FUNCTION_BLOCK "FB_ManInsp_V1.00"   // FB24, LAD
{ S7_Optimized_Access := 'TRUE' }
VERSION : 0.1
   VAR_INPUT
      IN_xCycleON : Bool;   // Cycle ON
      IN_xCycleONDel : Bool;   // Delayed cycle ON signal
      IN_xGeneralReset : Bool;   // General reset
      IN_xResetAlarms : Bool;   // Reset alarms
      IN_xFaultsEnabled : Bool;   // Faults enabled
      IN_dGlassBreakMachineIndex : DInt;   // Glass break machine index
      IN_dNumButtonDefect : DInt;   // Number of defect button
      IN_dNumQltDefect : DInt;   // Number of quality defect
      INPUT : Struct   // Digital inputs
         xPowerSupplyControl : Bool;   // L+.Power supply control
         xOpenRolls : Bool;   // SA.Open rolls
         xCloseRolls : Bool;   // SA.Close rolls
         rgxDefectButtons : Array[0..#CONST_MAX_DEFECT_BUTTONS_IND] of Bool;   // Defects buttons
         rgxQualityButtons : Array[0..#CONST_MAX_QUALITY_BUTTONS_IND] of Bool;   // Quality buttons
      END_STRUCT;
   END_VAR
   VAR_OUTPUT
      OUTPUT : Struct
         xFanCommand : Bool;   // Fan command
         xCloseRolls : Bool;   // YV.Close rolls
         xOpenRolls : Bool;   // YV.Open rolls
         xLampOpenCloseRolls : Bool;   // HL.Open/Close rolls
         rgxDefectButtonsLamp : Array[0..#CONST_MAX_DEFECT_BUTTONS_IND] of Bool;   // Defect buttons lamp
         rgxQualityButtonsLamp : Array[0..#CONST_MAX_QUALITY_BUTTONS_IND] of Bool;   // quality buttons lamp
      END_STRUCT;
   END_VAR
   VAR_IN_OUT
      INO_tFBAddDefect : "FB_Defects_Add_V1.00";   // Add defect DB
      INO_tOBInitialize : "GP_OB_Initialize";   // OB Initialize
      INO_tEncoder : "UDT_Encoder";   // Encoder data
      INO_tRibbon : "UDT_RibbonData";   // Ribbon data
      INO_xDefectBufferFull : Bool;   // Defect buffer full
   END_VAR
   VAR RETAIN
      tHMW : Struct   // HMI Write
         tMan : Struct   // Manual commands
            xFanCommand : Bool;   // Fan command {x|x|x|x|O}
            xSpare_1 : Bool;
            xSpare_2 : Bool;
            xSpare_3 : Bool;
            xSpare_4 : Bool;
            xSpare_5 : Bool;
            xSpare_6 : Bool;
            xSpare_7 : Bool;
            xSpare_8 : Bool;
            xSpare_9 : Bool;
            xSpare_10 : Bool;
            xSpare_11 : Bool;
            xSpare_12 : Bool;
            xSpare_13 : Bool;
            xSpare_14 : Bool;
            xSpare_15 : Bool;
         END_STRUCT;
         xEnDisManCom : Bool;   // Enable disable manual command {x|x|x|x|O}
         rgdButtonClass : Array[0..#CONST_MAX_DEFECT_BUTTONS_IND] of DInt;   // Buttons defect class {x|x|1|20|O}
         rgdButtonPosition_cmm : Array[0..#CONST_MAX_DEFECT_BUTTONS_IND] of DInt;   // Buttons defect position {mm/100|mm|-3000|3000|O}
         rgxEnabledContinuosDef : Array[0..#CONST_MAX_DEFECT_BUTTONS_IND] of Bool;   // Enable continuos defect {x|x|x|x|O}
         dDefectLength_cmm : DInt;   // Defect length [mm/100] {mm/100|mm|1|1000|O}
         dDefectWidth_cmm : DInt;   // Defect width [mm/100] {mm/100|mm|1|1000|O}
         dDistanceSnaproll_cmm : DInt;   // Distance from snaproll [mm/100] {mm/100|mm|1|70000|M}
         xUpdateDistanceSnaproll : Bool;   // Update distance from snaproll {x|x|x|x|M}
         dCalibDefectTheoPosX_cmm : DInt;   // Calibration. Theorical defect position X [mm/100] {mm/100|mm|1|7000|O}
         dCalibDefectRealPosX_cmm : DInt;   // Calibration. Real defect position X [mm/100] {mm/100|mm|1|7000|O}
         xDefectCalibration : Bool;   // Calibration.Calibrate defect {x|x|x|x|M}
      END_STRUCT;
      tHMR : Struct   // HMI Read
         xManComEn : Bool;   // Manual command enabled {x|x|x|x|O}
         dDistanceSnaproll_cmm : DInt;   // Distance from snaproll [mm/100] {mm/100|mm|x|x|M}
         tManFdbk : Struct   // Manual commands feedback
            xFanCommand : Bool;   // Fan command {x|x|x|x|O}
            xSpare_1 : Bool;
            xSpare_2 : Bool;
            xSpare_3 : Bool;
            xSpare_4 : Bool;
            xSpare_5 : Bool;
            xSpare_6 : Bool;
            xSpare_7 : Bool;
            xSpare_8 : Bool;
            xSpare_9 : Bool;
            xSpare_10 : Bool;
            xSpare_11 : Bool;
            xSpare_12 : Bool;
            xSpare_13 : Bool;
            xSpare_14 : Bool;
            xSpare_15 : Bool;
         END_STRUCT;
      END_STRUCT;
   END_VAR
   VAR
      tALM : Struct   // HMI Alarms
         tS : Struct   // Stopping faults machine
            xPowerSupplyControl : Bool;   // 1A222/1L+.Power supply control {X|X|X|X|O}
            xSpare_1 : Bool;
            xSpare_2 : Bool;
            xSpare_3 : Bool;
            xSpare_4 : Bool;
            xSpare_5 : Bool;
            xSpare_6 : Bool;
            xSpare_7 : Bool;
            xSpare_8 : Bool;
            xSpare_9 : Bool;
            xSpare_10 : Bool;
            xSpare_11 : Bool;
            xSpare_12 : Bool;
            xSpare_13 : Bool;
            xSpare_14 : Bool;
            xSpare_15 : Bool;
            xSpare_16 : Bool;
            xSpare_17 : Bool;
            xSpare_18 : Bool;
            xSpare_19 : Bool;
            xSpare_20 : Bool;
            xSpare_21 : Bool;
            xSpare_22 : Bool;
            xSpare_23 : Bool;
            xSpare_24 : Bool;
            xSpare_25 : Bool;
            xSpare_26 : Bool;
            xSpare_27 : Bool;
            xSpare_28 : Bool;
            xSpare_29 : Bool;
            xSpare_30 : Bool;
            xSpare_31 : Bool;
         END_STRUCT;
         tF : Struct   // Faults
            xSpare_0 : Bool;
            xSpare_1 : Bool;
            xSpare_2 : Bool;
            xSpare_3 : Bool;
            xSpare_4 : Bool;
            xSpare_5 : Bool;
            xSpare_6 : Bool;
            xSpare_7 : Bool;
            xSpare_8 : Bool;
            xSpare_9 : Bool;
            xSpare_10 : Bool;
            xSpare_11 : Bool;
            xSpare_12 : Bool;
            xSpare_13 : Bool;
            xSpare_14 : Bool;
            xSpare_15 : Bool;
            xSpare_16 : Bool;
            xSpare_17 : Bool;
            xSpare_18 : Bool;
            xSpare_19 : Bool;
            xSpare_20 : Bool;
            xSpare_21 : Bool;
            xSpare_22 : Bool;
            xSpare_23 : Bool;
            xSpare_24 : Bool;
            xSpare_25 : Bool;
            xSpare_26 : Bool;
            xSpare_27 : Bool;
            xSpare_28 : Bool;
            xSpare_29 : Bool;
            xSpare_30 : Bool;
            xSpare_31 : Bool;
         END_STRUCT;
         tW : Struct   // Warnings
            xSpare_0 : Bool;
            xSpare_1 : Bool;
            xSpare_2 : Bool;
            xSpare_3 : Bool;
            xSpare_4 : Bool;
            xSpare_5 : Bool;
            xSpare_6 : Bool;
            xSpare_7 : Bool;
            xSpare_8 : Bool;
            xSpare_9 : Bool;
            xSpare_10 : Bool;
            xSpare_11 : Bool;
            xSpare_12 : Bool;
            xSpare_13 : Bool;
            xSpare_14 : Bool;
            xSpare_15 : Bool;
            xSpare_16 : Bool;
            xSpare_17 : Bool;
            xSpare_18 : Bool;
            xSpare_19 : Bool;
            xSpare_20 : Bool;
            xSpare_21 : Bool;
            xSpare_22 : Bool;
            xSpare_23 : Bool;
            xSpare_24 : Bool;
            xSpare_25 : Bool;
            xSpare_26 : Bool;
            xSpare_27 : Bool;
            xSpare_28 : Bool;
            xSpare_29 : Bool;
            xSpare_30 : Bool;
            xSpare_31 : Bool;
         END_STRUCT;
      END_STRUCT;
      ST_xOutputEnable : Bool;   // Output enable
      ST_xCondOkMan : Bool;   // Condition ok manual command
      ST_xGlassBreak : Bool;   // Glass break under bridge
      ST_xStoppedFaults : Bool;   // Stopped faults
      ST_xFaults : Bool;   // Faults
      ST_xWarning : Bool;   // Warnings
      AUX_rgxDefectButtonsLast : Array[0..#CONST_MAX_DEFECT_BUTTONS_IND] of Bool;   // Last state of defect button
      AUX_rgxQualityButtonsLast : Array[0..#CONST_MAX_QUALITY_BUTTONS_IND] of Bool;   // Last state of quality buttons
      INO_tFBAddDefect1 : "FB_Defects_Add_V1.00";
      AUX_rgdLastInsDeftPos_cmm : Array[0..#CONST_MAX_DEFECT_BUTTONS_IND] of DInt;   // Last inserted defect position
   END_VAR
   VAR_TEMP
      TMP_dwValue : DWord;
      TMP_dIndex : DInt;
   END_VAR
   VAR CONSTANT
      CONST_DSTATUS_ANOMALY : DInt := 7;
      CONST_DSTATUS_RUN : DInt := 3;
      CONST_DSTATUS_IDLE : DInt := 1;
      CONST_DTIMEOUT_MS : DInt := 300000;   // Refill timeout [ms]
      CONST_MAX_DEFECT_BUTTONS : DInt := 16;   // Max defects buttons
      CONST_MAX_DEFECT_BUTTONS_IND : DInt := 15;   // Max defects buttons index (Always -1 than real)
      CONST_MAX_QUALITY_BUTTONS : DInt := 8;   // Max quality buttons
      CONST_MAX_QUALITY_BUTTONS_IND : DInt := 7;   // Max quality buttons index (Always -1 than real)
      CONST_MANUAL_DEFECT_SUBTYPE : DInt := 1000;   // Manual defect subtype
      CONST_QUALITY_DEFECT_CLASS : DInt := 21;   // Quality defect class
      CONST_QUALITY_SUBTYPE_EXACTPOS : DInt := 1001;   // Quality at exact position subtype
      CONST_CONTDEFLENGTH_CMM : DInt := 100000;   // Continuos defect length [mm/100]
      CONST_DBREAKUPOFF_CMM : DInt := 50000;   // Break upstream offset [mm/100]
      CONST_DBREAKDOWNOFF_CMM : DInt := 50000;   // Break downstream offset [mm/100]
   END_VAR
BEGIN

REGION Network 1: ####_CONSTANTS_####
END_REGION

REGION Network 2: ####_MATCH_####
END_REGION

REGION Network 3 (SCL): General reset
   IF #IN_xGeneralReset THEN

       FOR #TMP_dIndex := 0 TO #IN_dNumButtonDefect - 1 DO
           #tHMW.rgxEnabledContinuosDef[#TMP_dIndex] := FALSE;
       END_FOR;

   END_IF;
END_REGION

REGION Network 4: ####_HMI_LOGICS_####
END_REGION

REGION Network 5: Manual command enabled
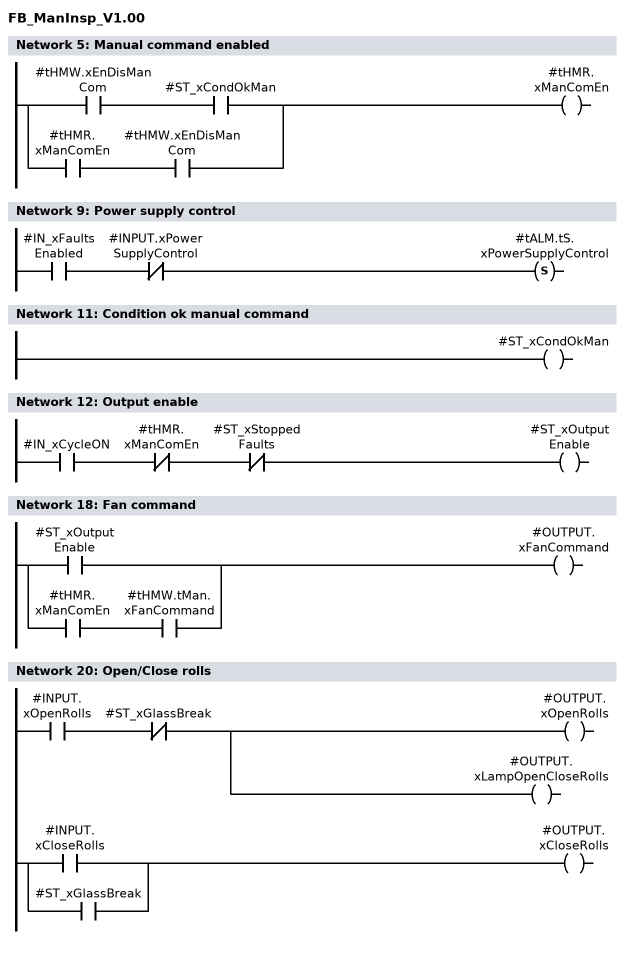
   RUNG wire#powerrail
      Contact( #tHMW.xEnDisManCom )
      Contact( #ST_xCondOkMan )
      wire#w1
      Coil( #tHMR.xManComEn )
   END_RUNG
   RUNG wire#powerrail
      Contact( #tHMR.xManComEn )
      Contact( #tHMW.xEnDisManCom )
   END_RUNG wire#w1
   // the same network as SCL:
   #tHMR.xManComEn := (#tHMW.xEnDisManCom AND #ST_xCondOkMan) OR (#tHMR.xManComEn AND #tHMW.xEnDisManCom);
END_REGION

REGION Network 6 (SCL): Manage HMI
   FOR #TMP_dIndex := 0 TO #IN_dNumButtonDefect - 1 DO

   (*    IF #tHMW.rgxEnableContinuosDef[#TMP_dIndex] THEN
           #tHMW.rgxEnableContinuosDef[#TMP_dIndex] := FALSE;
           #tHMR.rgxEnableContinuosDef[#TMP_dIndex] := TRUE;
           #AUX_rgdLastInsDeftPos_cmm[#TMP_dIndex] := #INO_tEncoder.dActualEncoderCounter_cmm;
       END_IF;

       IF #tHMW.rgxDisableContinuosDef[#TMP_dIndex] THEN
           #tHMW.rgxDisableContinuosDef[#TMP_dIndex] := FALSE;
           #tHMR.rgxEnableContinuosDef[#TMP_dIndex] := FALSE;
           #AUX_rgdLastInsDeftPos_cmm[#TMP_dIndex] := 0;

       END_IF; *)

       IF #tHMW.rgxEnabledContinuosDef[#TMP_dIndex] = true THEN
           #AUX_rgdLastInsDeftPos_cmm[#TMP_dIndex] := #INO_tEncoder.dActualEncoderCounter_cmm;
       ELSE
           #AUX_rgdLastInsDeftPos_cmm[#TMP_dIndex] := 0;
       END_IF;
   END_FOR;

   IF #tHMW.xUpdateDistanceSnaproll THEN
       #tHMW.xUpdateDistanceSnaproll := FALSE;
       #tHMR.dDistanceSnaproll_cmm := #tHMW.dDistanceSnaproll_cmm;
   END_IF;

   IF #tHMW.xDefectCalibration THEN
       #tHMW.xDefectCalibration := FALSE;
       #tHMR.dDistanceSnaproll_cmm += (#tHMW.dCalibDefectRealPosX_cmm - #tHMW.dCalibDefectTheoPosX_cmm);
   END_IF;
END_REGION

REGION Network 7: ####_ALARMS_####
END_REGION

REGION Network 8 (SCL): Reset alarms
   IF #IN_xResetAlarms THEN

       #TMP_dwValue := 0;

       SCATTER(IN:=#TMP_dwValue,
               OUT=>#tALM.tS);

       SCATTER(IN:=#TMP_dwValue,
               OUT=>#tALM.tF);

       SCATTER(IN:=#TMP_dwValue,
               OUT=>#tALM.tW);


   END_IF;
END_REGION

REGION Network 9: Power supply control
   RUNG wire#powerrail
      Contact( #IN_xFaultsEnabled )
      I_Contact( #INPUT.xPowerSupplyControl )
      S_Coil( #tALM.tS.xPowerSupplyControl )
   END_RUNG
   // the same network as SCL:
   IF #IN_xFaultsEnabled AND NOT #INPUT.xPowerSupplyControl THEN
       #tALM.tS.xPowerSupplyControl := TRUE;
   END_IF;
END_REGION

REGION Network 10: ####_STATUSES_####
END_REGION

REGION Network 11: Condition ok manual command
   RUNG wire#powerrail
      Coil( #ST_xCondOkMan )
   END_RUNG
   // the same network as SCL:
   #ST_xCondOkMan := TRUE;
END_REGION

REGION Network 12: Output enable
   RUNG wire#powerrail
      Contact( #IN_xCycleON )
      I_Contact( #tHMR.xManComEn )
      I_Contact( #ST_xStoppedFaults )
      Coil( #ST_xOutputEnable )
   END_RUNG
   // the same network as SCL:
   #ST_xOutputEnable := #IN_xCycleON AND NOT #tHMR.xManComEn AND NOT #ST_xStoppedFaults;
END_REGION

REGION Network 13 (SCL): Glass break calculation
   #INO_tRibbon.rgtGlassBreakRequest[#IN_dGlassBreakMachineIndex].IN_dDistanceSnaproll_cmm := #tHMR.dDistanceSnaproll_cmm;
   #INO_tRibbon.rgtGlassBreakRequest[#IN_dGlassBreakMachineIndex].IN_dDownstreamOffset_cmm := #CONST_DBREAKDOWNOFF_CMM;
   #INO_tRibbon.rgtGlassBreakRequest[#IN_dGlassBreakMachineIndex].IN_dUpstreamOffset_cmm := #CONST_DBREAKUPOFF_CMM;

   IF #INO_tRibbon.rgtGlassBreakRequest[#IN_dGlassBreakMachineIndex].OUT_xDataReady THEN
       #ST_xGlassBreak := #INO_tRibbon.rgtGlassBreakRequest[#IN_dGlassBreakMachineIndex].OUT_xGlassBreak;
   END_IF;

   IF #INO_tRibbon.rgtGlassBreakRequest[#IN_dGlassBreakMachineIndex].OUT_xDataReady OR NOT #INO_tRibbon.rgtGlassBreakRequest[#IN_dGlassBreakMachineIndex].IN_xRequestGlassBreak THEN
       #INO_tRibbon.rgtGlassBreakRequest[#IN_dGlassBreakMachineIndex].OUT_xDataReady := FALSE;
       #INO_tRibbon.rgtGlassBreakRequest[#IN_dGlassBreakMachineIndex].IN_xRequestGlassBreak := TRUE;
   END_IF;
END_REGION

REGION Network 14: ### PHASE AND LOGICS ###
END_REGION

REGION Network 15 (SCL): Manage pressed push button
   FOR #TMP_dIndex := 0 TO #IN_dNumQltDefect - 1 DO

       IF #INPUT.rgxQualityButtons[#TMP_dIndex] <> #AUX_rgxQualityButtonsLast[#TMP_dIndex] AND #INPUT.rgxQualityButtons[#TMP_dIndex]  = TRUE THEN

           #INO_tFBAddDefect(IN_dClass:=#CONST_QUALITY_DEFECT_CLASS,
              IN_dSubType:=#CONST_QUALITY_SUBTYPE_EXACTPOS,
              IN_dXPosition_cmm:=#INO_tEncoder.dActualEncoderCounter_cmm + #tHMR.dDistanceSnaproll_cmm,
              IN_dYPosition_cmm:=0,
              IN_dTotalLength_um:=1000,
              IN_dTotalWidth_um:=1000,
              IN_dCoreLength_um := 1000,
              IN_dCoreWidth_um:=1000,
              IN_dDistLength_um := 1000, 
              IN_dDistWidth_um:=1000,
              IN_dOptValue_mdptr:=0,
              OUT_xBufferFull => #INO_xDefectBufferFull,
              IN_strDefectID:='QUALITY_EXACT_POSITION');

       END_IF;

       #AUX_rgxQualityButtonsLast[#TMP_dIndex] := #INPUT.rgxQualityButtons[#TMP_dIndex];


   END_FOR;

   FOR #TMP_dIndex := 0 TO #IN_dNumButtonDefect - 1 DO

       IF #INPUT.rgxDefectButtons[#TMP_dIndex] <> #AUX_rgxDefectButtonsLast[#TMP_dIndex] AND #INPUT.rgxDefectButtons[#TMP_dIndex] THEN

           #INO_tFBAddDefect(IN_dClass:=#tHMW.rgdButtonClass[#TMP_dIndex],
              IN_dSubType:=#CONST_MANUAL_DEFECT_SUBTYPE,
              IN_dXPosition_cmm:=#INO_tEncoder.dActualEncoderCounter_cmm + #tHMR.dDistanceSnaproll_cmm,
              IN_dYPosition_cmm:=#tHMW.rgdButtonPosition_cmm[#TMP_dIndex],
              IN_dTotalLength_um:=#tHMW.dDefectLength_cmm * 10,
              IN_dTotalWidth_um:=#tHMW.dDefectWidth_cmm * 10,
              IN_dCoreLength_um := #tHMW.dDefectLength_cmm * 10,
              IN_dCoreWidth_um:=#tHMW.dDefectWidth_cmm * 10,
              IN_dDistLength_um := #tHMW.dDefectLength_cmm * 10,
              IN_dDistWidth_um:=#tHMW.dDefectWidth_cmm * 10,
              IN_dOptValue_mdptr:=0,
              OUT_xBufferFull => #INO_xDefectBufferFull,
              IN_strDefectID:='MANUAL_DEFECT');

       END_IF;

       #AUX_rgxDefectButtonsLast[#TMP_dIndex] := #INPUT.rgxDefectButtons[#TMP_dIndex];

       IF ((#INO_tEncoder.dActualEncoderCounter_cmm - #AUX_rgdLastInsDeftPos_cmm[#TMP_dIndex]) >= 0) AND (#tHMW.rgxEnabledContinuosDef[#TMP_dIndex]) THEN

           #INO_tFBAddDefect(IN_dClass:=#tHMW.rgdButtonClass[#TMP_dIndex],
              IN_dSubType:=#CONST_MANUAL_DEFECT_SUBTYPE,
              IN_dXPosition_cmm:=#INO_tEncoder.dActualEncoderCounter_cmm + #tHMR.dDistanceSnaproll_cmm,
              IN_dYPosition_cmm:=#tHMW.rgdButtonPosition_cmm[#TMP_dIndex],
              IN_dTotalLength_um:=#CONST_CONTDEFLENGTH_CMM * 10,
              IN_dTotalWidth_um:=#tHMW.dDefectWidth_cmm * 10,
              IN_dCoreLength_um :=#CONST_CONTDEFLENGTH_CMM * 10,
              IN_dCoreWidth_um:=#tHMW.dDefectWidth_cmm * 10,
              IN_dDistLength_um := #CONST_CONTDEFLENGTH_CMM * 10,
              IN_dDistWidth_um:=#tHMW.dDefectWidth_cmm * 10,
              IN_dOptValue_mdptr:=0,
              OUT_xBufferFull => #INO_xDefectBufferFull,
              IN_strDefectID:='MANUAL_DEFECT');

               #AUX_rgdLastInsDeftPos_cmm[#TMP_dIndex] += #CONST_CONTDEFLENGTH_CMM;

       END_IF;

   END_FOR;
END_REGION

REGION Network 16 (SCL): ### HMI STATUS ###
   #tHMR.tManFdbk.xFanCommand := #OUTPUT.xFanCommand AND #tHMW.tMan.xFanCommand;
END_REGION

REGION Network 17: ####_OUTPUT_####
END_REGION

REGION Network 18: Fan command
   RUNG wire#powerrail
      Contact( #ST_xOutputEnable )
      wire#w1
      Coil( #OUTPUT.xFanCommand )
   END_RUNG
   RUNG wire#powerrail
      Contact( #tHMR.xManComEn )
      Contact( #tHMW.tMan.xFanCommand )
   END_RUNG wire#w1
   // the same network as SCL:
   #OUTPUT.xFanCommand := #ST_xOutputEnable OR (#tHMR.xManComEn AND #tHMW.tMan.xFanCommand);
END_REGION

REGION Network 19 (SCL): Lamp output
   FOR #TMP_dIndex := 0 TO #IN_dNumButtonDefect - 1 DO
       #OUTPUT.rgxDefectButtonsLamp[#TMP_dIndex] := #INPUT.rgxDefectButtons[#TMP_dIndex];
   END_FOR;

   FOR #TMP_dIndex := 0 TO #IN_dNumQltDefect - 1 DO
       #OUTPUT.rgxQualityButtonsLamp[#TMP_dIndex] := #INPUT.rgxQualityButtons[#TMP_dIndex];
   END_FOR;
END_REGION

REGION Network 20: Open/Close rolls
   RUNG wire#powerrail
      Contact( #INPUT.xOpenRolls )
      I_Contact( #ST_xGlassBreak )
      wire#w1
      Coil( #OUTPUT.xOpenRolls )
   END_RUNG
   RUNG wire#w1
      Coil( #OUTPUT.xLampOpenCloseRolls )
   END_RUNG
   RUNG wire#powerrail
      Contact( #INPUT.xCloseRolls )
      wire#w2
      Coil( #OUTPUT.xCloseRolls )
   END_RUNG
   RUNG wire#powerrail
      Contact( #ST_xGlassBreak )
   END_RUNG wire#w2
   // the same network as SCL:
   #OUTPUT.xOpenRolls := #INPUT.xOpenRolls AND NOT #ST_xGlassBreak;
   #OUTPUT.xLampOpenCloseRolls := #OUTPUT.xOpenRolls;
   #OUTPUT.xCloseRolls := #INPUT.xCloseRolls OR #ST_xGlassBreak;
END_REGION
END_FUNCTION_BLOCK

// folder: 03_Programs_Logics/MCC1200/25_WanderCamera

FUNCTION_BLOCK "FB_WanderCamera_V1.00"   // FB22, LAD
{ S7_Optimized_Access := 'TRUE' }
VERSION : 0.1
   VAR_INPUT
      IN_xCycleON : Bool;   // Cycle ON
      IN_xCycleONDel : Bool;   // Delayed cycle ON signal
      IN_xGeneralReset : Bool;   // General reset
      IN_xResetAlarms : Bool;   // Reset alarms
      IN_xFaultsEnabled : Bool;   // Faults enabled
      IN_tInterfaceID : Hw_Any;   // Interface ID
      IN_tID : Conn_Ouc;   // Connection ID
      IN_tRemoteAddress : IP_V4;   // Remote IP address
      IN_uiRemotePort : UInt;   // Remote port
      IN_dGlassBreakMachineIndex : DInt;   // Glass break machine index
      IN_dGlassDataMachineIndex : DInt;   // Glass data machine index
   END_VAR
   VAR_IN_OUT
      INO_tTrack : "UDT_CapData_Tracking";   // Tracking plate
      INO_tRibbon : "UDT_RibbonData";   // Ribbon data
   END_VAR
   VAR RETAIN
      tHMR : Struct
         dCameraStatus : DInt := 0;   // Camera status (1=Disabled, 3=Enabled, 7=Anomaly) {x|x|x|x|O}
         dDistanceFromSnaproll_cmm : DInt := 0;   // Distance from snaproll [mm/100] {mm/100|mm|x|x|O}
         dCurrentGrossWidth_cmm : DInt := 0;   // Current gross width [mm/100] {mm/100|mm|x|x|O}
         dCurrentNetWidth_cmm : DInt := 0;   // Current net width [mm/100] {mm/100|mm|x|x|O}
         dCurrentGrossWander_cmm : DInt := 0;   // Current gross wander [mm/100] {mm/100|mm|x|x|O}
         dCurrentNetWander_cmm : DInt := 0;   // Current net wander [mm/100] {mm/100|mm|x|x|O}
      END_STRUCT;
      tHMW : Struct
         dDistanceFromSnaproll_cmm : DInt := 0;   // Distance from snaproll [mm/100] {mm/100|mm|0|30000|M}
         xUpdateDistanceFromSnaproll : Bool := 0;   // Update distance from snaproll {x|x|x|x|M}
      END_STRUCT;
   END_VAR
   VAR
      tALM : Struct   // HMI Alarms
         tS : Struct   // Stopping faults
            xCameraNotConnected : Bool;   // Camera system not connected
            xSendError : Bool;   // Sending data error
            xSendTimeout : Bool;   // Sending data timeout
            xRecvTimeout : Bool;   // Receiving data timeout
            xWanderOutLimits : Bool;   // Wander outside limits
            xCameraInError : Bool;   // Camera system in error
            xSpare_6 : Bool;
            xSpare_7 : Bool;
            xSpare_8 : Bool;
            xSpare_9 : Bool;
            xSpare_10 : Bool;
            xSpare_11 : Bool;
            xSpare_12 : Bool;
            xSpare_13 : Bool;
            xSpare_14 : Bool;
            xSpare_15 : Bool;
            xSpare_16 : Bool;
            xSpare_17 : Bool;
            xSpare_18 : Bool;
            xSpare_19 : Bool;
            xSpare_20 : Bool;
            xSpare_21 : Bool;
            xSpare_22 : Bool;
            xSpare_23 : Bool;
            xSpare_24 : Bool;
            xSpare_25 : Bool;
            xSpare_26 : Bool;
            xSpare_27 : Bool;
            xSpare_28 : Bool;
            xSpare_29 : Bool;
            xSpare_30 : Bool;
            xSpare_31 : Bool;
         END_STRUCT;
         tF : Struct   // Faults
            xSpare_0 : Bool;
            xSpare_1 : Bool;
            xSpare_2 : Bool;
            xSpare_3 : Bool;
            xSpare_4 : Bool;
            xSpare_5 : Bool;
            xSpare_6 : Bool;
            xSpare_7 : Bool;
            xSpare_8 : Bool;
            xSpare_9 : Bool;
            xSpare_10 : Bool;
            xSpare_11 : Bool;
            xSpare_12 : Bool;
            xSpare_13 : Bool;
            xSpare_14 : Bool;
            xSpare_15 : Bool;
            xSpare_16 : Bool;
            xSpare_17 : Bool;
            xSpare_18 : Bool;
            xSpare_19 : Bool;
            xSpare_20 : Bool;
            xSpare_21 : Bool;
            xSpare_22 : Bool;
            xSpare_23 : Bool;
            xSpare_24 : Bool;
            xSpare_25 : Bool;
            xSpare_26 : Bool;
            xSpare_27 : Bool;
            xSpare_28 : Bool;
            xSpare_29 : Bool;
            xSpare_30 : Bool;
            xSpare_31 : Bool;
         END_STRUCT;
         tW : Struct   // Warnings
            xSpare_0 : Bool;
            xSpare_1 : Bool;
            xSpare_2 : Bool;
            xSpare_3 : Bool;
            xSpare_4 : Bool;
            xSpare_5 : Bool;
            xSpare_6 : Bool;
            xSpare_7 : Bool;
            xSpare_8 : Bool;
            xSpare_9 : Bool;
            xSpare_10 : Bool;
            xSpare_11 : Bool;
            xSpare_12 : Bool;
            xSpare_13 : Bool;
            xSpare_14 : Bool;
            xSpare_15 : Bool;
            xSpare_16 : Bool;
            xSpare_17 : Bool;
            xSpare_18 : Bool;
            xSpare_19 : Bool;
            xSpare_20 : Bool;
            xSpare_21 : Bool;
            xSpare_22 : Bool;
            xSpare_23 : Bool;
            xSpare_24 : Bool;
            xSpare_25 : Bool;
            xSpare_26 : Bool;
            xSpare_27 : Bool;
            xSpare_28 : Bool;
            xSpare_29 : Bool;
            xSpare_30 : Bool;
            xSpare_31 : Bool;
         END_STRUCT;
      END_STRUCT;
      ST_xStoppingFaults : Bool;   // Stopping faults
      ST_xFaults : Bool;   // Faults
      ST_xOuputEnable : Bool;   // Output enable
      ST_xCondOkMan : Bool;   // Condition ok manual command
      ST_xPhaseProgr : Bool;   // Phase in progress
      ST_xWarnings : Bool;   // Warnings
      ST_xGlassBreak : Bool;   // Glass break
      ST_xWandOutLimits : Bool;   // Wander out of limits
      OS_xNewDataAvailable : Bool;   // New data received from camera
      tPhases : Struct   // Phases
         xSendTelegram : Bool;   // Send telegram
         xEndSendTelegram : Bool;   // End send telegram
         xSpare2 : Bool;
         xSpare3 : Bool;
         xSpare4 : Bool;
         xSpare5 : Bool;
         xSpare6 : Bool;
         xSpare7 : Bool;
         xSpare8 : Bool;
         xSpare9 : Bool;
         xSpare10 : Bool;
         xSpare11 : Bool;
         xSpare12 : Bool;
         xSpare13 : Bool;
         xSpare14 : Bool;
         xSpare15 : Bool;
         xSpare16 : Bool;
         xSpare17 : Bool;
         xSpare18 : Bool;
         xSpare19 : Bool;
         xSpare20 : Bool;
         xSpare21 : Bool;
         xSpare22 : Bool;
         xSpare23 : Bool;
         xSpare24 : Bool;
         xSpare25 : Bool;
         xSpare26 : Bool;
         xSpare27 : Bool;
         xSpare28 : Bool;
         xSpare29 : Bool;
         xSpare30 : Bool;
         xSpare31 : Bool;
      END_STRUCT;
      FB_TSend : TSEND_C;
      FB_TReceive : TRCV_C;
      AUX_tConnData : TCON_IP_v4;   // Connection data structure
      AUX_xResetSendConnection : Bool;   // Reset the estabilished send connection
      AUX_xResetRecvConnection : Bool;   // Reset the estabilished receive connection
      AUX_dNumByteToSend : DInt;   // Number of byte to send
      AUX_rdtTempRecvBuffer : Array[0..55] of Byte;   // Temporary receive buffer
      AUX_rdtRecvBuffer : Struct   // Receive buffer
         dLung : DInt := 0;   // Record length
         dID : DInt := 0;   // Incremental packet number
         dTime1 : DInt := 0;   // Timing #1
         dTime2 : DInt := 0;   // Timing #2
         dStato : DInt := 0;   // Wander status (0=Not in measure, 1=in measure, 2=in calibration)
         dGrossZeroSide_um : DInt := 0;   // Gross zero side [um]
         dNetExtZeroSide_um : DInt := 0;   // Net ext. zero side [um]
         dNetCenterZeroSide_um : DInt := 0;   // Net center zero side [um]
         dNetZeroSide_um : DInt := 0;   // Net zero side [um]
         dGrossOppSide_um : DInt := 0;   // Gross opposite side [um]
         dNetExtOppoSide_um : DInt := 0;   // Net ext. opposite side [um]
         dNetCenterOppoSide_um : DInt := 0;   // Net center opposite side [um]
         dNetOppoSide_um : DInt := 0;   // Net opposite side [um]
         dLength : DInt := 0;   // Record length
      END_STRUCT;
      AUX_rgtSendBuffer : Struct   // Send buffer
         dLung : DInt;   // Packet lenght
         dID : DInt;   // ID Message
         dThick_um : DInt;   // Thickness [um]
      END_STRUCT;
      AUX_rgtSendBuffer_LittleEndian : Array[0..11] of Byte;   // Send buffer
      tmON_TimeoutRecvData : TON_TIME;   // Timeout receive data
      tmON_TimeoutSendData : TON_TIME;   // Timeout sending data
      tmON_SendData : TON_TIME;   // Timer TON send data
   END_VAR
   VAR_TEMP
      TMP_xPrepareTelegram : Bool;
      TMP_dPos : DInt;
      TMP_dwValue : DWord;
      TMP_iRetVal : Int;
   END_VAR
   VAR CONSTANT
      CONST_BCONNTYPE : Byte := 16#0B;   // Connection type
      CONST_DTIMEOUTSENDDATA_MS : DInt := 5000;   // Timeout sending data [ms]
      CONST_DTIMEOUTNEWDATA_MS : DInt := 60000;   // Timeout receive new data [ms]
      CONST_DTIMESENDDATA_MS : DInt := 2000;   // Time send data [ms]
   END_VAR
   VAR_TEMP   // added for the SCL form of the ladder/FBD networks
      _w1 : Bool;
   END_VAR
BEGIN

REGION Network 1: ####_COSTANTS_####
END_REGION

REGION Network 2: ####_MATCH_####
END_REGION

REGION Network 3: ####_ALARMS_####
END_REGION

REGION Network 4 (SCL): Reset alarms
   IF #IN_xResetAlarms THEN

       #TMP_dwValue := 0;

       SCATTER(IN:=#TMP_dwValue,
               OUT=>#tALM.tS);

       SCATTER(IN:=#TMP_dwValue,
               OUT=>#tALM.tF);

       SCATTER(IN:=#TMP_dwValue,
               OUT=>#tALM.tW);


   END_IF;
END_REGION

REGION Network 5: Camera system not connected
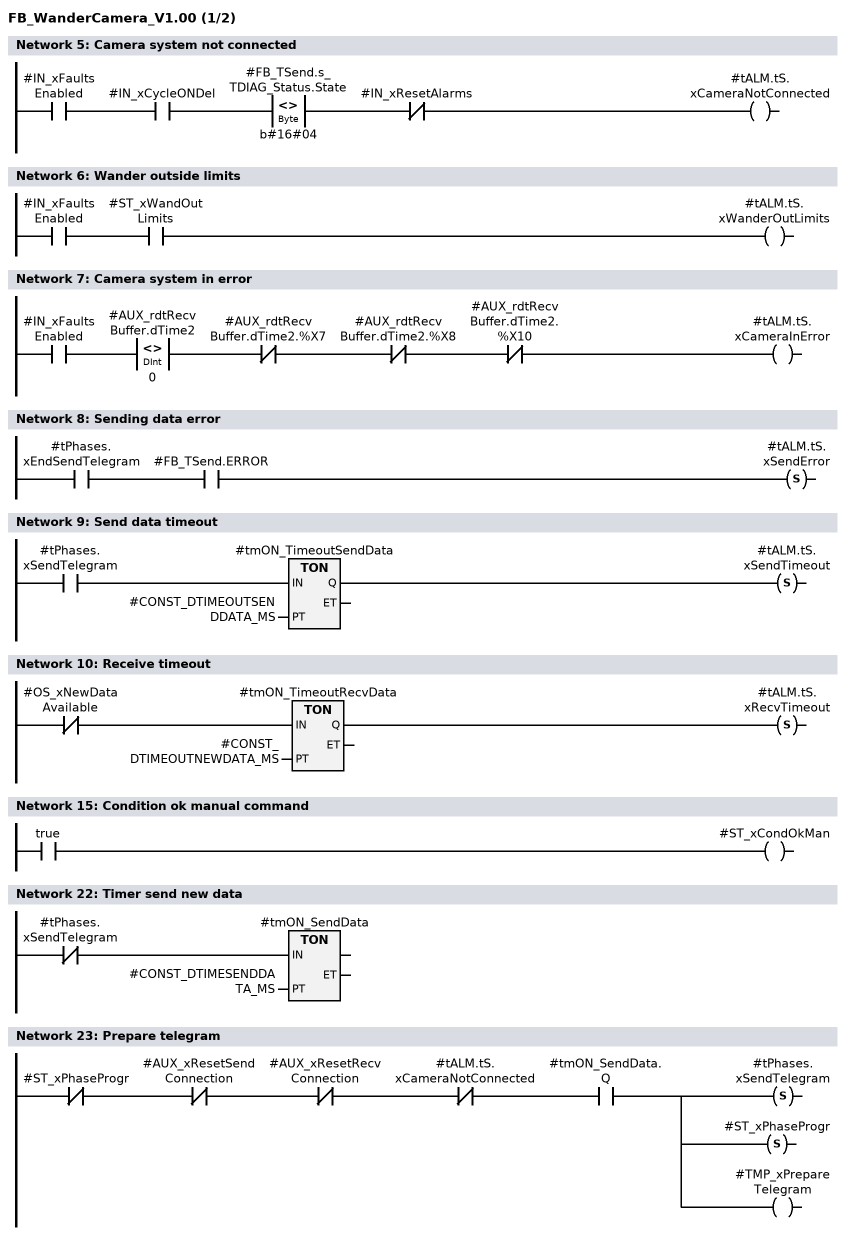
   RUNG wire#powerrail
      Contact( #IN_xFaultsEnabled )
      Contact( #IN_xCycleONDel )
      { S7_Templates := "SrcType := Byte" } NE_Contact(in1 := #FB_TSend.s_TDIAG_Status.State, in2 := b#16#04)
      I_Contact( #IN_xResetAlarms )
      Coil( #tALM.tS.xCameraNotConnected )
   END_RUNG
   // the same network as SCL:
   #tALM.tS.xCameraNotConnected := #IN_xFaultsEnabled AND #IN_xCycleONDel AND (#FB_TSend.s_TDIAG_Status.State <> b#16#04) AND NOT #IN_xResetAlarms;
END_REGION

REGION Network 6: Wander outside limits
   RUNG wire#powerrail
      Contact( #IN_xFaultsEnabled )
      Contact( #ST_xWandOutLimits )
      Coil( #tALM.tS.xWanderOutLimits )
   END_RUNG
   // the same network as SCL:
   #tALM.tS.xWanderOutLimits := #IN_xFaultsEnabled AND #ST_xWandOutLimits;
END_REGION

REGION Network 7: Camera system in error
   RUNG wire#powerrail
      Contact( #IN_xFaultsEnabled )
      { S7_Templates := "SrcType := DInt" } NE_Contact(in1 := #AUX_rdtRecvBuffer.dTime2, in2 := 0)
      I_Contact( #AUX_rdtRecvBuffer.dTime2.%X7 )
      I_Contact( #AUX_rdtRecvBuffer.dTime2.%X8 )
      I_Contact( #AUX_rdtRecvBuffer.dTime2.%X10 )
      Coil( #tALM.tS.xCameraInError )
   END_RUNG
   // the same network as SCL:
   #tALM.tS.xCameraInError := #IN_xFaultsEnabled AND (#AUX_rdtRecvBuffer.dTime2 <> 0) AND NOT #AUX_rdtRecvBuffer.dTime2.%X7 AND NOT #AUX_rdtRecvBuffer.dTime2.%X8 AND NOT #AUX_rdtRecvBuffer.dTime2.%X10;
END_REGION

REGION Network 8: Sending data error
   RUNG wire#powerrail
      Contact( #tPhases.xEndSendTelegram )
      Contact( #FB_TSend.ERROR )
      S_Coil( #tALM.tS.xSendError )
   END_RUNG
   // the same network as SCL:
   IF #tPhases.xEndSendTelegram AND #FB_TSend.ERROR THEN #tALM.tS.xSendError := TRUE; END_IF;
END_REGION

REGION Network 9: Send data timeout
   #tmON_TimeoutSendData(IN := #tPhases.xSendTelegram, PT := #CONST_DTIMEOUTSENDDATA_MS);   // TON
   IF #tmON_TimeoutSendData.Q THEN #tALM.tS.xSendTimeout := TRUE; END_IF;
END_REGION

REGION Network 10: Receive timeout
   #tmON_TimeoutRecvData(IN := NOT #OS_xNewDataAvailable, PT := #CONST_DTIMEOUTNEWDATA_MS);   // TON
   IF #tmON_TimeoutRecvData.Q THEN #tALM.tS.xRecvTimeout := TRUE; END_IF;
END_REGION

REGION Network 11 (SCL): Calculate general statuses
   GATHER(IN:=#tALM.tS,
          OUT=>#TMP_dwValue);

   IF #TMP_dwValue <> 0 THEN
       #ST_xStoppingFaults := TRUE;
   ELSE
       #ST_xStoppingFaults := FALSE;
   END_IF;

   GATHER(IN:=#tALM.tF,
          OUT=>#TMP_dwValue);

   IF #TMP_dwValue <> 0 THEN
       #ST_xFaults := TRUE;
   ELSE
       #ST_xFaults := FALSE;
   END_IF;

   GATHER(IN:=#tALM.tW,
          OUT=>#TMP_dwValue);

   IF #TMP_dwValue <> 0 THEN
       #ST_xWarnings := TRUE;
   ELSE
       #ST_xWarnings := FALSE;
   END_IF;
END_REGION

REGION Network 12: ####_HMI_LOGICS_####
END_REGION

REGION Network 13 (SCL): Manage HMI request

   REGION Distance from snaproll calibration

       IF #tHMW.xUpdateDistanceFromSnaproll THEN

           #tHMR.dDistanceFromSnaproll_cmm := #tHMW.dDistanceFromSnaproll_cmm;

           #tHMW.xUpdateDistanceFromSnaproll  := FALSE;

       END_IF;

   END_REGION
END_REGION

REGION Network 14: ####_STATUSES_####
END_REGION

REGION Network 15: Condition ok manual command
   RUNG wire#powerrail
      Contact( true )
      Coil( #ST_xCondOkMan )
   END_RUNG
   // the same network as SCL:
   #ST_xCondOkMan := true;
END_REGION

REGION Network 16: ####_PHASES_&_LOGICS_####
END_REGION

REGION Network 17 (SCL): Glass break calculation
   #INO_tRibbon.rgtGlassBreakRequest[#IN_dGlassBreakMachineIndex].IN_dDistanceSnaproll_cmm := #tHMR.dDistanceFromSnaproll_cmm;
   #INO_tRibbon.rgtGlassBreakRequest[#IN_dGlassBreakMachineIndex].IN_dDownstreamOffset_cmm := 0;
   #INO_tRibbon.rgtGlassBreakRequest[#IN_dGlassBreakMachineIndex].IN_dUpstreamOffset_cmm := 0;

   IF #INO_tRibbon.rgtGlassBreakRequest[#IN_dGlassBreakMachineIndex].OUT_xDataReady THEN
       #ST_xGlassBreak := #INO_tRibbon.rgtGlassBreakRequest[#IN_dGlassBreakMachineIndex].OUT_xGlassBreak;
   END_IF;

   IF #INO_tRibbon.rgtGlassBreakRequest[#IN_dGlassBreakMachineIndex].OUT_xDataReady OR NOT #INO_tRibbon.rgtGlassBreakRequest[#IN_dGlassBreakMachineIndex].IN_xRequestGlassBreak THEN
       #INO_tRibbon.rgtGlassBreakRequest[#IN_dGlassBreakMachineIndex].OUT_xDataReady := FALSE;
       #INO_tRibbon.rgtGlassBreakRequest[#IN_dGlassBreakMachineIndex].IN_xRequestGlassBreak := TRUE;
   END_IF;
END_REGION

REGION Network 18 (SCL): Normalize data
   IF NOT (#ST_xGlassBreak) THEN
       #tHMR.dCurrentGrossWidth_cmm := ((#AUX_rdtRecvBuffer.dGrossZeroSide_um * -1) + #AUX_rdtRecvBuffer.dGrossOppSide_um) / 10;
       #tHMR.dCurrentNetWidth_cmm := ((#AUX_rdtRecvBuffer.dNetZeroSide_um * -1) + #AUX_rdtRecvBuffer.dNetOppoSide_um) / 10;

       #tHMR.dCurrentGrossWander_cmm := (#tHMR.dCurrentGrossWidth_cmm / 2) - ((#AUX_rdtRecvBuffer.dGrossZeroSide_um * -1) / 10);
       #tHMR.dCurrentNetWander_cmm := (#tHMR.dCurrentNetWidth_cmm / 2) - ((#AUX_rdtRecvBuffer.dNetZeroSide_um * -1) / 10);

       //Check the limits
       #ST_xWandOutLimits := 0;

       IF #tHMR.dCurrentGrossWidth_cmm > "DMAXGROSSWIDTH_CMM" THEN

           #ST_xWandOutLimits := 1;

       END_IF;

       IF #tHMR.dCurrentGrossWidth_cmm < "DMINGROSSWIDTH_CMM" THEN

           #ST_xWandOutLimits := 1;

       END_IF;

       IF #tHMR.dCurrentNetWidth_cmm > "DMAXNETWIDTH_CMM" THEN

           #ST_xWandOutLimits := 1;

       END_IF;

       IF #tHMR.dCurrentNetWidth_cmm < "DMINNETWIDTH_CMM" THEN

           #ST_xWandOutLimits := 1;

       END_IF;

       IF #tHMR.dCurrentGrossWander_cmm > "DMAXGROSSWANDER_CMM" THEN

           #ST_xWandOutLimits := 1;

       END_IF;

       IF #tHMR.dCurrentGrossWander_cmm < "DMINGROSSWANDER_CMM" THEN

           #ST_xWandOutLimits := 1;

       END_IF;

       IF #tHMR.dCurrentNetWander_cmm > "DMAXNETWANDER_CMM" THEN

           #ST_xWandOutLimits := 1;

       END_IF;

       IF #tHMR.dCurrentNetWander_cmm < "DMINNETWANDER_CMM" THEN

           #ST_xWandOutLimits := 1;

       END_IF;
   END_IF;
END_REGION

REGION Network 19 (SCL): ####_HMI_STATUSES_####
   IF #ST_xStoppingFaults THEN
       #tHMR.dCameraStatus := 7;
   ELSE
       #tHMR.dCameraStatus := 3;
   END_IF;
END_REGION

REGION Network 20: ####_ETHERNET_TO_CAMERA_####
END_REGION

REGION Network 21 (SCL): Initialize connection data
   IF #IN_xGeneralReset  THEN

       #AUX_tConnData.InterfaceId := #IN_tInterfaceID;
       #AUX_tConnData.ID := #IN_tID;
       #AUX_tConnData.ConnectionType := #CONST_BCONNTYPE;
       #AUX_tConnData.ActiveEstablished := FALSE;
       #AUX_tConnData.RemotePort := 0;
       #AUX_tConnData.LocalPort := #IN_uiRemotePort;

       //Reset della fasi
       #TMP_dwValue := 0;
       SCATTER(IN:=#TMP_dwValue,
               OUT=>#tPhases);



   END_IF;

   #AUX_xResetRecvConnection := #IN_xGeneralReset;
   #AUX_xResetSendConnection := #IN_xGeneralReset;
END_REGION

REGION Network 22: Timer send new data
   #tmON_SendData(IN := NOT #tPhases.xSendTelegram, PT := #CONST_DTIMESENDDATA_MS);   // TON
END_REGION

REGION Network 23: Prepare telegram
   RUNG wire#powerrail
      I_Contact( #ST_xPhaseProgr )
      I_Contact( #AUX_xResetSendConnection )
      I_Contact( #AUX_xResetRecvConnection )
      I_Contact( #tALM.tS.xCameraNotConnected )
      Contact( #tmON_SendData.Q )
      wire#w1
      S_Coil( #tPhases.xSendTelegram )
   END_RUNG
   RUNG wire#w1
      S_Coil( #ST_xPhaseProgr )
   END_RUNG
   RUNG wire#w1
      Coil( #TMP_xPrepareTelegram )
   END_RUNG
   // the same network as SCL:
   #_w1 := NOT #ST_xPhaseProgr AND NOT #AUX_xResetSendConnection AND NOT #AUX_xResetRecvConnection AND NOT #tALM.tS.xCameraNotConnected AND #tmON_SendData.Q;
   IF #_w1 THEN
       #tPhases.xSendTelegram := TRUE;
       #ST_xPhaseProgr := TRUE;
   END_IF;
   #TMP_xPrepareTelegram := #_w1;
END_REGION

REGION Network 24 (SCL): Prepare telegram
   IF #TMP_xPrepareTelegram THEN